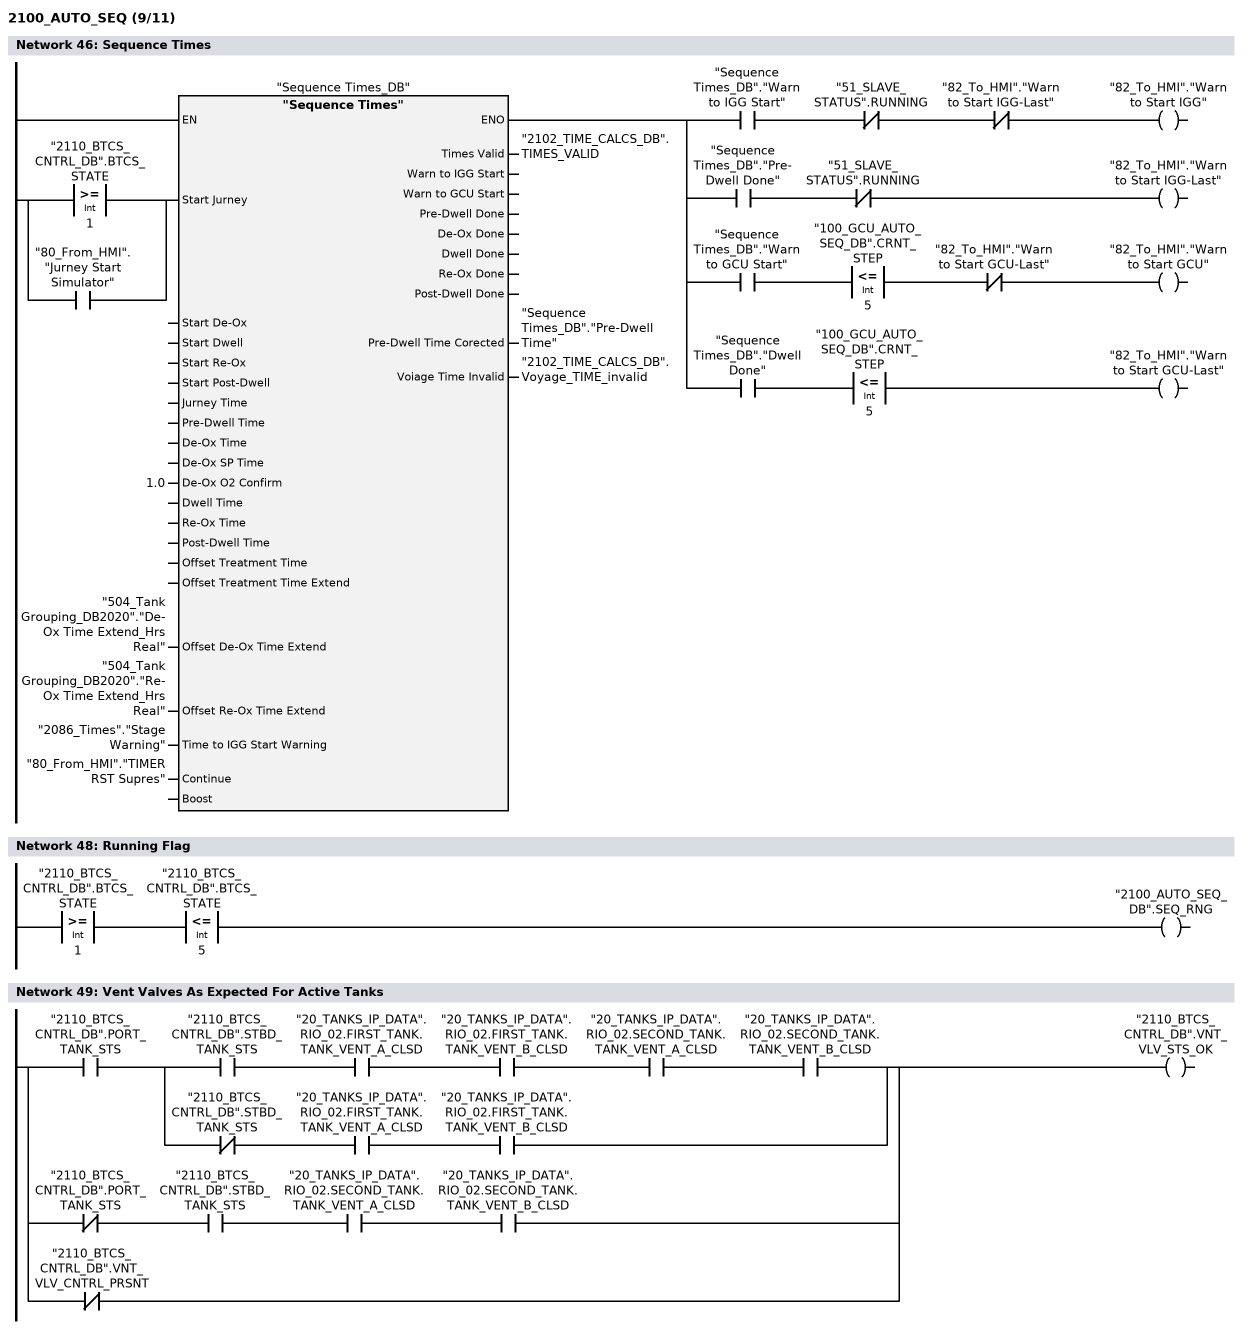
   RUNG wire#powerrail
      "Sequence Times_DB"("Start Jurney" := wire#w1, "Start De-Ox" :=, "Start Dwell" :=, "Start Re-Ox" :=, "Start Post-Dwell" :=, "Jurney Time" :=, "Pre-Dwell Time" :=, "De-Ox Time" :=, "De-Ox SP Time" :=, "De-Ox O2 Confirm" := 1.0, "Dwell Time" :=, "Re-Ox Time" :=, "Post-Dwell Time" :=, "Offset Treatment Time" :=, "Offset Treatment Time Extend" :=, "Offset De-Ox Time Extend" := "504_Tank Grouping_DB2020"."De-Ox Time Extend_Hrs Real", "Offset Re-Ox Time Extend" := "504_Tank Grouping_DB2020"."Re-Ox Time Extend_Hrs Real", "Time to IGG Start Warning" := "2086_Times"."Stage Warning", Continue := "80_From_HMI"."TIMER RST Supres", Boost :=, "Times Valid" => "2102_TIME_CALCS_DB".TIMES_VALID, "Warn to IGG Start" =>, "Warn to GCU Start" =>, "Pre-Dwell Done" =>, "De-Ox Done" =>, "Dwell Done" =>, "Re-Ox Done" =>, "Post-Dwell Done" =>, "Pre-Dwell Time Corected" => "Sequence Times_DB"."Pre-Dwell Time", "Voiage Time Invalid" => "2102_TIME_CALCS_DB".Voyage_TIME_invalid)
      wire#w2
      Contact( "Sequence Times_DB"."Warn to IGG Start" )
      I_Contact( "51_SLAVE_STATUS".RUNNING )
      I_Contact( "82_To_HMI"."Warn to Start IGG-Last" )
      Coil( "82_To_HMI"."Warn to Start IGG" )
   END_RUNG
   RUNG wire#powerrail
      { S7_Templates := "SrcType := Int" } GE_Contact(in1 := "2110_BTCS_CNTRL_DB".BTCS_STATE, in2 := 1)
   END_RUNG wire#w1
   RUNG wire#powerrail
      Contact( "80_From_HMI"."Jurney Start Simulator" )
   END_RUNG wire#w1
   RUNG wire#w2
      Contact( "Sequence Times_DB"."Pre-Dwell Done" )
      I_Contact( "51_SLAVE_STATUS".RUNNING )
      Coil( "82_To_HMI"."Warn to Start IGG-Last" )
   END_RUNG
   RUNG wire#w2
      Contact( "Sequence Times_DB"."Warn to GCU Start" )
      { S7_Templates := "SrcType := Int" } LE_Contact(in1 := "100_GCU_AUTO_SEQ_DB".CRNT_STEP, in2 := 5)
      I_Contact( "82_To_HMI"."Warn to Start GCU-Last" )
      Coil( "82_To_HMI"."Warn to Start GCU" )
   END_RUNG
   RUNG wire#w2
      Contact( "Sequence Times_DB"."Dwell Done" )
      { S7_Templates := "SrcType := Int" } LE_Contact(in1 := "100_GCU_AUTO_SEQ_DB".CRNT_STEP, in2 := 5)
      Coil( "82_To_HMI"."Warn to Start GCU-Last" )
   END_RUNG
   // the same network as SCL:
   "Sequence Times_DB"("Start Jurney" := ("2110_BTCS_CNTRL_DB".BTCS_STATE >= 1) OR "80_From_HMI"."Jurney Start Simulator",   // "Sequence Times"
                       "De-Ox O2 Confirm" := 1.0,
                       "Offset De-Ox Time Extend" := "504_Tank Grouping_DB2020"."De-Ox Time Extend_Hrs Real",
                       "Offset Re-Ox Time Extend" := "504_Tank Grouping_DB2020"."Re-Ox Time Extend_Hrs Real",
                       "Time to IGG Start Warning" := "2086_Times"."Stage Warning",
                       Continue := "80_From_HMI"."TIMER RST Supres",
                       "Times Valid" => "2102_TIME_CALCS_DB".TIMES_VALID,
                       "Pre-Dwell Time Corected" => "Sequence Times_DB"."Pre-Dwell Time",
                       "Voiage Time Invalid" => "2102_TIME_CALCS_DB".Voyage_TIME_invalid,
                       ENO => #_w1);
   "82_To_HMI"."Warn to Start IGG" := #_w1 AND "Sequence Times_DB"."Warn to IGG Start" AND NOT "51_SLAVE_STATUS".RUNNING AND NOT "82_To_HMI"."Warn to Start IGG-Last";
   "82_To_HMI"."Warn to Start IGG-Last" := #_w1 AND "Sequence Times_DB"."Pre-Dwell Done" AND NOT "51_SLAVE_STATUS".RUNNING;
   "82_To_HMI"."Warn to Start GCU" := #_w1 AND "Sequence Times_DB"."Warn to GCU Start" AND ("100_GCU_AUTO_SEQ_DB".CRNT_STEP <= 5) AND NOT "82_To_HMI"."Warn to Start GCU-Last";
   "82_To_HMI"."Warn to Start GCU-Last" := #_w1 AND "Sequence Times_DB"."Dwell Done" AND ("100_GCU_AUTO_SEQ_DB".CRNT_STEP <= 5);
END_REGION

REGION Network 48: Running Flag
   RUNG wire#powerrail
      { S7_Templates := "SrcType := Int" } GE_Contact(in1 := "2110_BTCS_CNTRL_DB".BTCS_STATE, in2 := 1)
      { S7_Templates := "SrcType := Int" } LE_Contact(in1 := "2110_BTCS_CNTRL_DB".BTCS_STATE, in2 := 5)
      Coil( "2100_AUTO_SEQ_DB".SEQ_RNG )
   END_RUNG
   // the same network as SCL:
   "2100_AUTO_SEQ_DB".SEQ_RNG := ("2110_BTCS_CNTRL_DB".BTCS_STATE >= 1) AND ("2110_BTCS_CNTRL_DB".BTCS_STATE <= 5);
END_REGION

REGION Network 49: Vent Valves As Expected For Active Tanks
   RUNG wire#powerrail
      Contact( "2110_BTCS_CNTRL_DB".PORT_TANK_STS )
      wire#w1
      Contact( "2110_BTCS_CNTRL_DB".STBD_TANK_STS )
      Contact( "20_TANKS_IP_DATA".RIO_02.FIRST_TANK.TANK_VENT_A_CLSD )
      Contact( "20_TANKS_IP_DATA".RIO_02.FIRST_TANK.TANK_VENT_B_CLSD )
      Contact( "20_TANKS_IP_DATA".RIO_02.SECOND_TANK.TANK_VENT_A_CLSD )
      Contact( "20_TANKS_IP_DATA".RIO_02.SECOND_TANK.TANK_VENT_B_CLSD )
      wire#w2
      Coil( "2110_BTCS_CNTRL_DB".VNT_VLV_STS_OK )
   END_RUNG
   RUNG wire#w1
      I_Contact( "2110_BTCS_CNTRL_DB".STBD_TANK_STS )
      Contact( "20_TANKS_IP_DATA".RIO_02.FIRST_TANK.TANK_VENT_A_CLSD )
      Contact( "20_TANKS_IP_DATA".RIO_02.FIRST_TANK.TANK_VENT_B_CLSD )
   END_RUNG wire#w2
   RUNG wire#powerrail
      I_Contact( "2110_BTCS_CNTRL_DB".PORT_TANK_STS )
      Contact( "2110_BTCS_CNTRL_DB".STBD_TANK_STS )
      Contact( "20_TANKS_IP_DATA".RIO_02.SECOND_TANK.TANK_VENT_A_CLSD )
      Contact( "20_TANKS_IP_DATA".RIO_02.SECOND_TANK.TANK_VENT_B_CLSD )
   END_RUNG wire#w2
   RUNG wire#powerrail
      I_Contact( "2110_BTCS_CNTRL_DB".VNT_VLV_CNTRL_PRSNT )
   END_RUNG wire#w2
   // the same network as SCL:
   "2110_BTCS_CNTRL_DB".VNT_VLV_STS_OK := ("2110_BTCS_CNTRL_DB".PORT_TANK_STS AND (("2110_BTCS_CNTRL_DB".STBD_TANK_STS AND "20_TANKS_IP_DATA".RIO_02.FIRST_TANK.TANK_VENT_A_CLSD AND "20_TANKS_IP_DATA".RIO_02.FIRST_TANK.TANK_VENT_B_CLSD AND "20_TANKS_IP_DATA".RIO_02.SECOND_TANK.TANK_VENT_A_CLSD AND "20_TANKS_IP_DATA".RIO_02.SECOND_TANK.TANK_VENT_B_CLSD) OR (NOT "2110_BTCS_CNTRL_DB".STBD_TANK_STS AND "20_TANKS_IP_DATA".RIO_02.FIRST_TANK.TANK_VENT_A_CLSD AND "20_TANKS_IP_DATA".RIO_02.FIRST_TANK.TANK_VENT_B_CLSD))) OR (NOT "2110_BTCS_CNTRL_DB".PORT_TANK_STS AND "2110_BTCS_CNTRL_DB".STBD_TANK_STS AND "20_TANKS_IP_DATA".RIO_02.SECOND_TANK.TANK_VENT_A_CLSD AND "20_TANKS_IP_DATA".RIO_02.SECOND_TANK.TANK_VENT_B_CLSD) OR NOT "2110_BTCS_CNTRL_DB".VNT_VLV_CNTRL_PRSNT;
END_REGION

REGION Network 50: GTT Valves As Expected For Active Tanks (condition used from Tank Grouping FB)
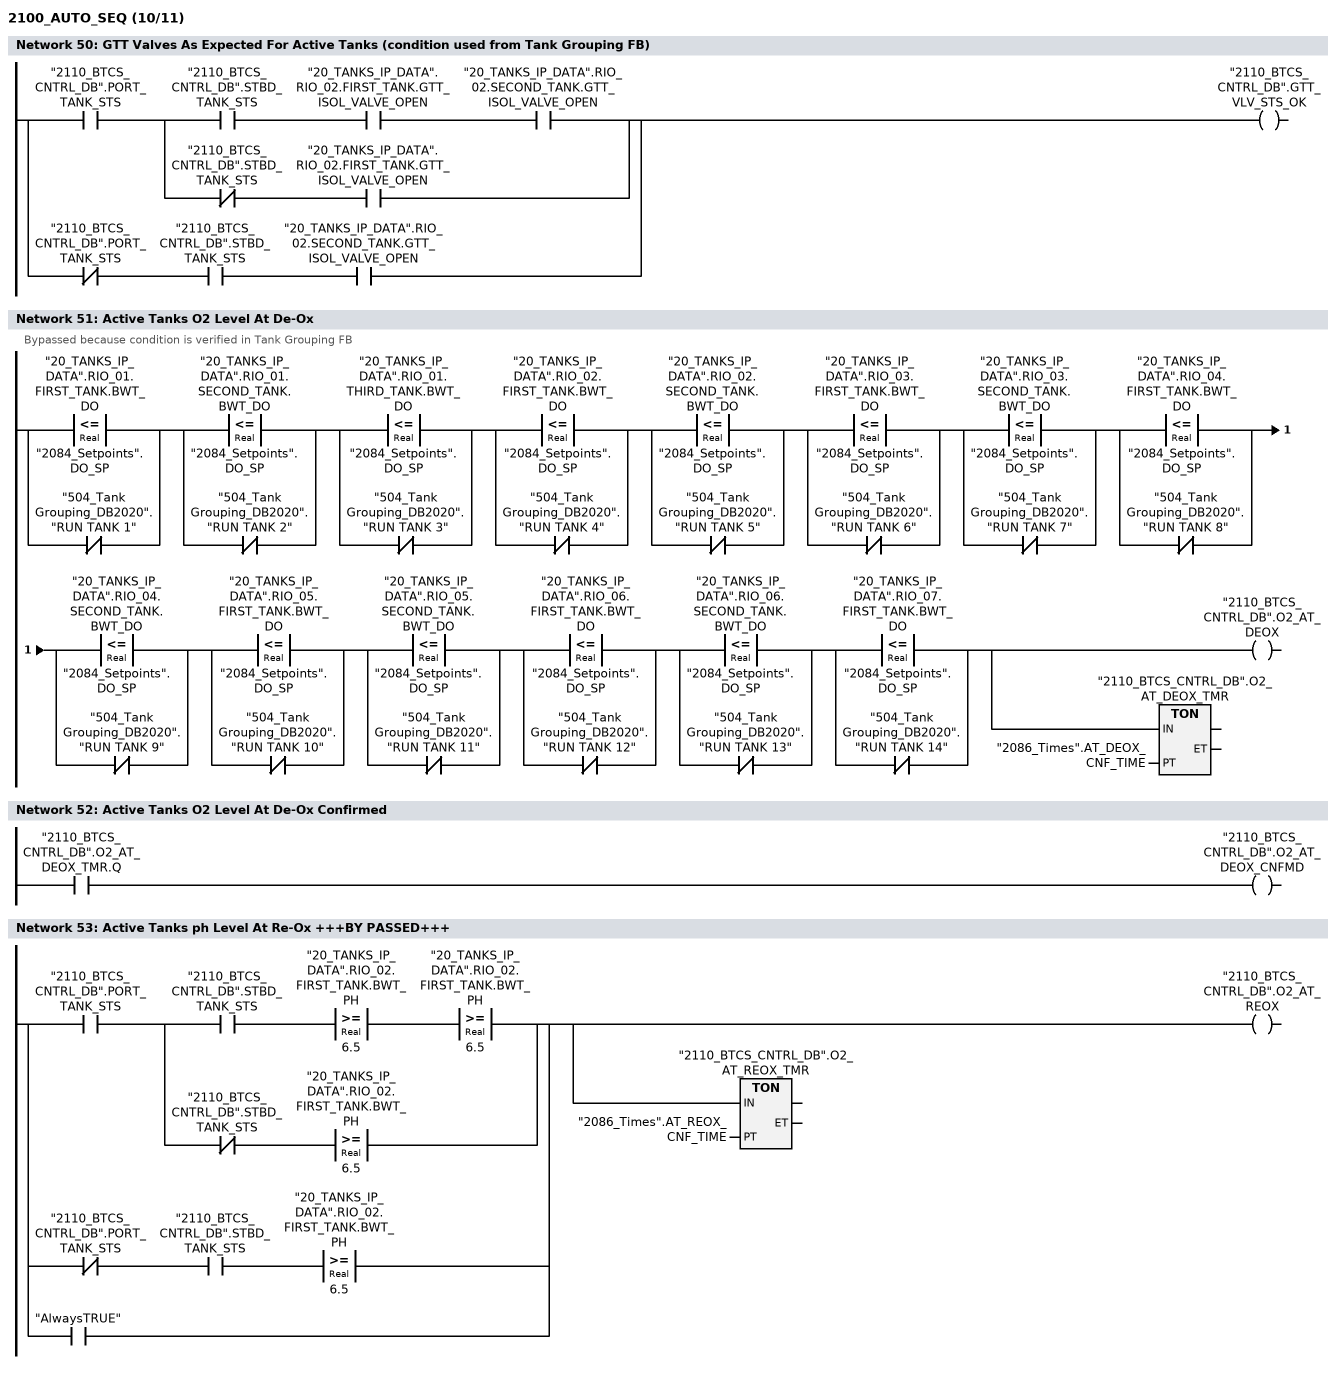
   RUNG wire#powerrail
      Contact( "2110_BTCS_CNTRL_DB".PORT_TANK_STS )
      wire#w1
      Contact( "2110_BTCS_CNTRL_DB".STBD_TANK_STS )
      Contact( "20_TANKS_IP_DATA".RIO_02.FIRST_TANK.GTT_ISOL_VALVE_OPEN )
      Contact( "20_TANKS_IP_DATA".RIO_02.SECOND_TANK.GTT_ISOL_VALVE_OPEN )
      wire#w2
      Coil( "2110_BTCS_CNTRL_DB".GTT_VLV_STS_OK )
   END_RUNG
   RUNG wire#w1
      I_Contact( "2110_BTCS_CNTRL_DB".STBD_TANK_STS )
      Contact( "20_TANKS_IP_DATA".RIO_02.FIRST_TANK.GTT_ISOL_VALVE_OPEN )
   END_RUNG wire#w2
   RUNG wire#powerrail
      I_Contact( "2110_BTCS_CNTRL_DB".PORT_TANK_STS )
      Contact( "2110_BTCS_CNTRL_DB".STBD_TANK_STS )
      Contact( "20_TANKS_IP_DATA".RIO_02.SECOND_TANK.GTT_ISOL_VALVE_OPEN )
   END_RUNG wire#w2
   // the same network as SCL:
   "2110_BTCS_CNTRL_DB".GTT_VLV_STS_OK := ("2110_BTCS_CNTRL_DB".PORT_TANK_STS AND (("2110_BTCS_CNTRL_DB".STBD_TANK_STS AND "20_TANKS_IP_DATA".RIO_02.FIRST_TANK.GTT_ISOL_VALVE_OPEN AND "20_TANKS_IP_DATA".RIO_02.SECOND_TANK.GTT_ISOL_VALVE_OPEN) OR (NOT "2110_BTCS_CNTRL_DB".STBD_TANK_STS AND "20_TANKS_IP_DATA".RIO_02.FIRST_TANK.GTT_ISOL_VALVE_OPEN))) OR (NOT "2110_BTCS_CNTRL_DB".PORT_TANK_STS AND "2110_BTCS_CNTRL_DB".STBD_TANK_STS AND "20_TANKS_IP_DATA".RIO_02.SECOND_TANK.GTT_ISOL_VALVE_OPEN);
END_REGION

REGION Network 51: Active Tanks O2 Level At De-Ox
   // Bypassed because condition is verified in Tank Grouping FB
   "2110_BTCS_CNTRL_DB".O2_AT_DEOX := (("20_TANKS_IP_DATA".RIO_01.FIRST_TANK.BWT_DO <= "2084_Setpoints".DO_SP) OR NOT "504_Tank Grouping_DB2020"."RUN TANK 1") AND (("20_TANKS_IP_DATA".RIO_01.SECOND_TANK.BWT_DO <= "2084_Setpoints".DO_SP) OR NOT "504_Tank Grouping_DB2020"."RUN TANK 2") AND (("20_TANKS_IP_DATA".RIO_01.THIRD_TANK.BWT_DO <= "2084_Setpoints".DO_SP) OR NOT "504_Tank Grouping_DB2020"."RUN TANK 3") AND (("20_TANKS_IP_DATA".RIO_02.FIRST_TANK.BWT_DO <= "2084_Setpoints".DO_SP) OR NOT "504_Tank Grouping_DB2020"."RUN TANK 4") AND (("20_TANKS_IP_DATA".RIO_02.SECOND_TANK.BWT_DO <= "2084_Setpoints".DO_SP) OR NOT "504_Tank Grouping_DB2020"."RUN TANK 5") AND (("20_TANKS_IP_DATA".RIO_03.FIRST_TANK.BWT_DO <= "2084_Setpoints".DO_SP) OR NOT "504_Tank Grouping_DB2020"."RUN TANK 6") AND (("20_TANKS_IP_DATA".RIO_03.SECOND_TANK.BWT_DO <= "2084_Setpoints".DO_SP) OR NOT "504_Tank Grouping_DB2020"."RUN TANK 7") AND (("20_TANKS_IP_DATA".RIO_04.FIRST_TANK.BWT_DO <= "2084_Setpoints".DO_SP) OR NOT "504_Tank Grouping_DB2020"."RUN TANK 8") AND (("20_TANKS_IP_DATA".RIO_04.SECOND_TANK.BWT_DO <= "2084_Setpoints".DO_SP) OR NOT "504_Tank Grouping_DB2020"."RUN TANK 9") AND (("20_TANKS_IP_DATA".RIO_05.FIRST_TANK.BWT_DO <= "2084_Setpoints".DO_SP) OR NOT "504_Tank Grouping_DB2020"."RUN TANK 10") AND (("20_TANKS_IP_DATA".RIO_05.SECOND_TANK.BWT_DO <= "2084_Setpoints".DO_SP) OR NOT "504_Tank Grouping_DB2020"."RUN TANK 11") AND (("20_TANKS_IP_DATA".RIO_06.FIRST_TANK.BWT_DO <= "2084_Setpoints".DO_SP) OR NOT "504_Tank Grouping_DB2020"."RUN TANK 12") AND (("20_TANKS_IP_DATA".RIO_06.SECOND_TANK.BWT_DO <= "2084_Setpoints".DO_SP) OR NOT "504_Tank Grouping_DB2020"."RUN TANK 13") AND (("20_TANKS_IP_DATA".RIO_07.FIRST_TANK.BWT_DO <= "2084_Setpoints".DO_SP) OR NOT "504_Tank Grouping_DB2020"."RUN TANK 14");
   "2110_BTCS_CNTRL_DB".O2_AT_DEOX_TMR.TON(IN := "2110_BTCS_CNTRL_DB".O2_AT_DEOX,
                           PT := "2086_Times".AT_DEOX_CNF_TIME);
END_REGION

REGION Network 52: Active Tanks O2 Level At De-Ox Confirmed
   RUNG wire#powerrail
      Contact( "2110_BTCS_CNTRL_DB".O2_AT_DEOX_TMR.Q )
      Coil( "2110_BTCS_CNTRL_DB".O2_AT_DEOX_CNFMD )
   END_RUNG
   // the same network as SCL:
   "2110_BTCS_CNTRL_DB".O2_AT_DEOX_CNFMD := "2110_BTCS_CNTRL_DB".O2_AT_DEOX_TMR.Q;
END_REGION

REGION Network 53: Active Tanks ph Level At Re-Ox +++BY PASSED+++
   "2110_BTCS_CNTRL_DB".O2_AT_REOX := ("2110_BTCS_CNTRL_DB".PORT_TANK_STS AND (("2110_BTCS_CNTRL_DB".STBD_TANK_STS AND ("20_TANKS_IP_DATA".RIO_02.FIRST_TANK.BWT_PH >= 6.5) AND ("20_TANKS_IP_DATA".RIO_02.FIRST_TANK.BWT_PH >= 6.5)) OR (NOT "2110_BTCS_CNTRL_DB".STBD_TANK_STS AND ("20_TANKS_IP_DATA".RIO_02.FIRST_TANK.BWT_PH >= 6.5)))) OR (NOT "2110_BTCS_CNTRL_DB".PORT_TANK_STS AND "2110_BTCS_CNTRL_DB".STBD_TANK_STS AND ("20_TANKS_IP_DATA".RIO_02.FIRST_TANK.BWT_PH >= 6.5)) OR "AlwaysTRUE";
   "2110_BTCS_CNTRL_DB".O2_AT_REOX_TMR.TON(IN := "2110_BTCS_CNTRL_DB".O2_AT_REOX,
                           PT := "2086_Times".AT_REOX_CNF_TIME);
END_REGION

REGION Network 54: Active Tanks ph Level At Re-Ox Confirmed
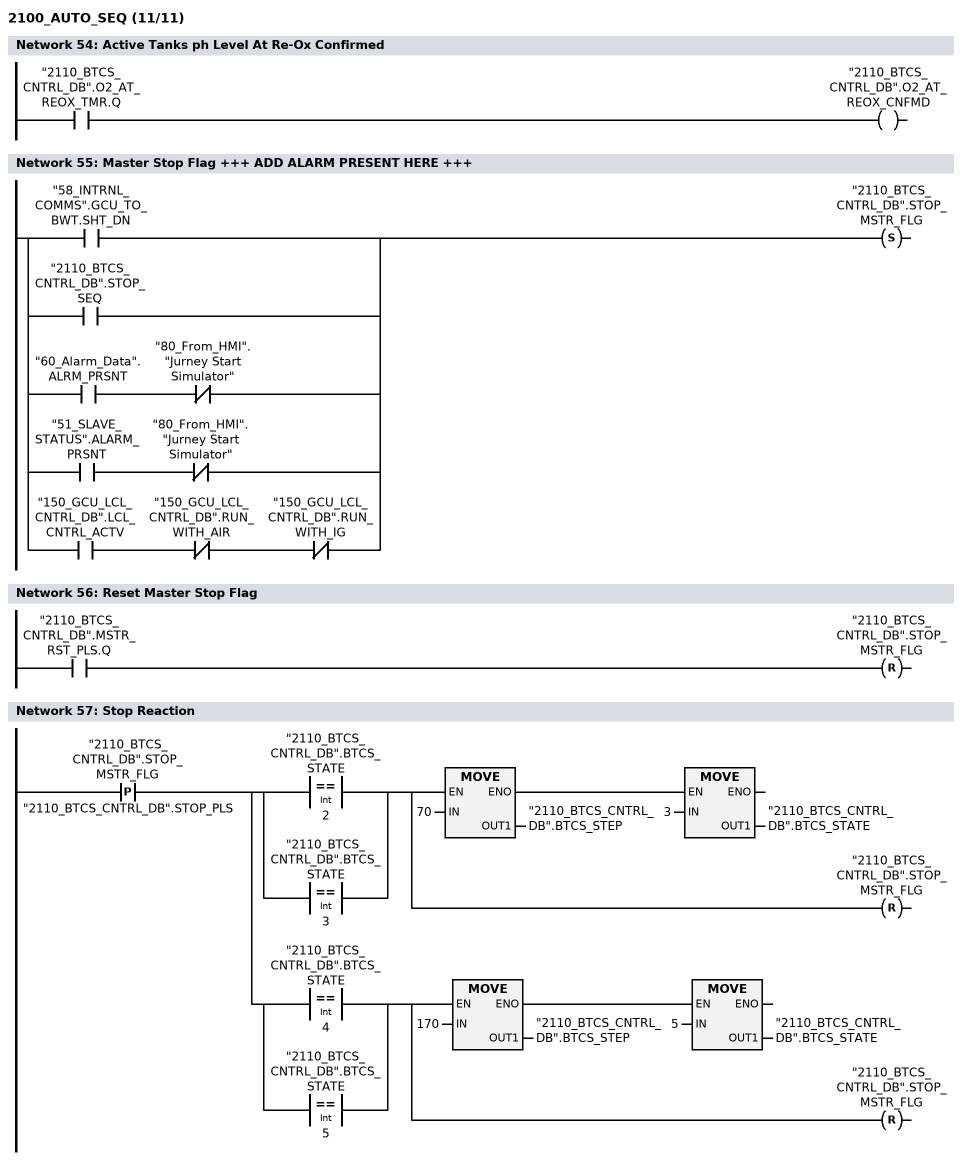
   RUNG wire#powerrail
      Contact( "2110_BTCS_CNTRL_DB".O2_AT_REOX_TMR.Q )
      Coil( "2110_BTCS_CNTRL_DB".O2_AT_REOX_CNFMD )
   END_RUNG
   // the same network as SCL:
   "2110_BTCS_CNTRL_DB".O2_AT_REOX_CNFMD := "2110_BTCS_CNTRL_DB".O2_AT_REOX_TMR.Q;
END_REGION

REGION Network 55: Master Stop Flag +++ ADD ALARM PRESENT HERE +++
   RUNG wire#powerrail
      Contact( "58_INTRNL_COMMS".GCU_TO_BWT.SHT_DN )
      wire#w1
      S_Coil( "2110_BTCS_CNTRL_DB".STOP_MSTR_FLG )
   END_RUNG
   RUNG wire#powerrail
      Contact( "2110_BTCS_CNTRL_DB".STOP_SEQ )
   END_RUNG wire#w1
   RUNG wire#powerrail
      Contact( "60_Alarm_Data".ALRM_PRSNT )
      I_Contact( "80_From_HMI"."Jurney Start Simulator" )
   END_RUNG wire#w1
   RUNG wire#powerrail
      Contact( "51_SLAVE_STATUS".ALARM_PRSNT )
      I_Contact( "80_From_HMI"."Jurney Start Simulator" )
   END_RUNG wire#w1
   RUNG wire#powerrail
      Contact( "150_GCU_LCL_CNTRL_DB".LCL_CNTRL_ACTV )
      I_Contact( "150_GCU_LCL_CNTRL_DB".RUN_WITH_AIR )
      I_Contact( "150_GCU_LCL_CNTRL_DB".RUN_WITH_IG )
   END_RUNG wire#w1
   // the same network as SCL:
   IF "58_INTRNL_COMMS".GCU_TO_BWT.SHT_DN OR "2110_BTCS_CNTRL_DB".STOP_SEQ OR ("60_Alarm_Data".ALRM_PRSNT AND NOT "80_From_HMI"."Jurney Start Simulator") OR ("51_SLAVE_STATUS".ALARM_PRSNT AND NOT "80_From_HMI"."Jurney Start Simulator") OR ("150_GCU_LCL_CNTRL_DB".LCL_CNTRL_ACTV AND NOT "150_GCU_LCL_CNTRL_DB".RUN_WITH_AIR AND NOT "150_GCU_LCL_CNTRL_DB".RUN_WITH_IG) THEN
       "2110_BTCS_CNTRL_DB".STOP_MSTR_FLG := TRUE;
   END_IF;
END_REGION

REGION Network 56: Reset Master Stop Flag
   RUNG wire#powerrail
      Contact( "2110_BTCS_CNTRL_DB".MSTR_RST_PLS.Q )
      R_Coil( "2110_BTCS_CNTRL_DB".STOP_MSTR_FLG )
   END_RUNG
   // the same network as SCL:
   IF "2110_BTCS_CNTRL_DB".MSTR_RST_PLS.Q THEN "2110_BTCS_CNTRL_DB".STOP_MSTR_FLG := FALSE; END_IF;
END_REGION

REGION Network 57: Stop Reaction
   RUNG wire#powerrail
      P_Contact(operand := "2110_BTCS_CNTRL_DB".STOP_MSTR_FLG, bit := "2110_BTCS_CNTRL_DB".STOP_PLS)
      wire#w1
      { S7_Templates := "SrcType := Int" } EQ_Contact(in1 := "2110_BTCS_CNTRL_DB".BTCS_STATE, in2 := 2)
      wire#w2
      Move(in := 70, out1 => "2110_BTCS_CNTRL_DB".BTCS_STEP)
      Move(in := 3, out1 => "2110_BTCS_CNTRL_DB".BTCS_STATE)
   END_RUNG
   RUNG wire#w1
      { S7_Templates := "SrcType := Int" } EQ_Contact(in1 := "2110_BTCS_CNTRL_DB".BTCS_STATE, in2 := 3)
   END_RUNG wire#w2
   RUNG wire#w2
      R_Coil( "2110_BTCS_CNTRL_DB".STOP_MSTR_FLG )
   END_RUNG
   RUNG wire#w1
      { S7_Templates := "SrcType := Int" } EQ_Contact(in1 := "2110_BTCS_CNTRL_DB".BTCS_STATE, in2 := 4)
      wire#w3
      Move(in := 170, out1 => "2110_BTCS_CNTRL_DB".BTCS_STEP)
      Move(in := 5, out1 => "2110_BTCS_CNTRL_DB".BTCS_STATE)
   END_RUNG
   RUNG wire#w1
      { S7_Templates := "SrcType := Int" } EQ_Contact(in1 := "2110_BTCS_CNTRL_DB".BTCS_STATE, in2 := 5)
   END_RUNG wire#w3
   RUNG wire#w3
      R_Coil( "2110_BTCS_CNTRL_DB".STOP_MSTR_FLG )
   END_RUNG
   // the same network as SCL:
   #_w1 := "2110_BTCS_CNTRL_DB".STOP_MSTR_FLG AND NOT "2110_BTCS_CNTRL_DB".STOP_PLS;   // rising edge of "2110_BTCS_CNTRL_DB".STOP_MSTR_FLG
   "2110_BTCS_CNTRL_DB".STOP_PLS := "2110_BTCS_CNTRL_DB".STOP_MSTR_FLG;
   IF #_w1 AND (("2110_BTCS_CNTRL_DB".BTCS_STATE = 2) OR ("2110_BTCS_CNTRL_DB".BTCS_STATE = 3)) THEN
       "2110_BTCS_CNTRL_DB".BTCS_STEP := 70;
   END_IF;
   #_w2 := #_w1 AND (("2110_BTCS_CNTRL_DB".BTCS_STATE = 2) OR ("2110_BTCS_CNTRL_DB".BTCS_STATE = 3));
   IF #_w2 THEN
       "2110_BTCS_CNTRL_DB".BTCS_STATE := 3;
       "2110_BTCS_CNTRL_DB".STOP_MSTR_FLG := FALSE;
   END_IF;
   IF #_w1 AND (("2110_BTCS_CNTRL_DB".BTCS_STATE = 4) OR ("2110_BTCS_CNTRL_DB".BTCS_STATE = 5)) THEN
       "2110_BTCS_CNTRL_DB".BTCS_STEP := 170;
   END_IF;
   #_w3 := #_w1 AND (("2110_BTCS_CNTRL_DB".BTCS_STATE = 4) OR ("2110_BTCS_CNTRL_DB".BTCS_STATE = 5));
   IF #_w3 THEN
       "2110_BTCS_CNTRL_DB".BTCS_STATE := 5;
       "2110_BTCS_CNTRL_DB".STOP_MSTR_FLG := FALSE;
   END_IF;
END_REGION
END_FUNCTION

FUNCTION "2102_TIME_CALCS" : Void   // FC2102, LAD
TITLE = Time Calculations
{ S7_Optimized_Access := 'TRUE' }
AUTHOR : JRS
VERSION : 0.1
// For calculating time periods associated with the BTCS
   VAR_TEMP
      T_REAL : Real;
   END_VAR
   VAR_TEMP   // added for the SCL form of the ladder/FBD networks
      _w1 : Bool;
      _w2 : Bool;
      _w3 : Bool;
      _w4 : Bool;
      _w5 : Bool;
      _w6 : Bool;
      _w7 : Bool;
   END_VAR
BEGIN

REGION Network 2: Minutes Phase Difference
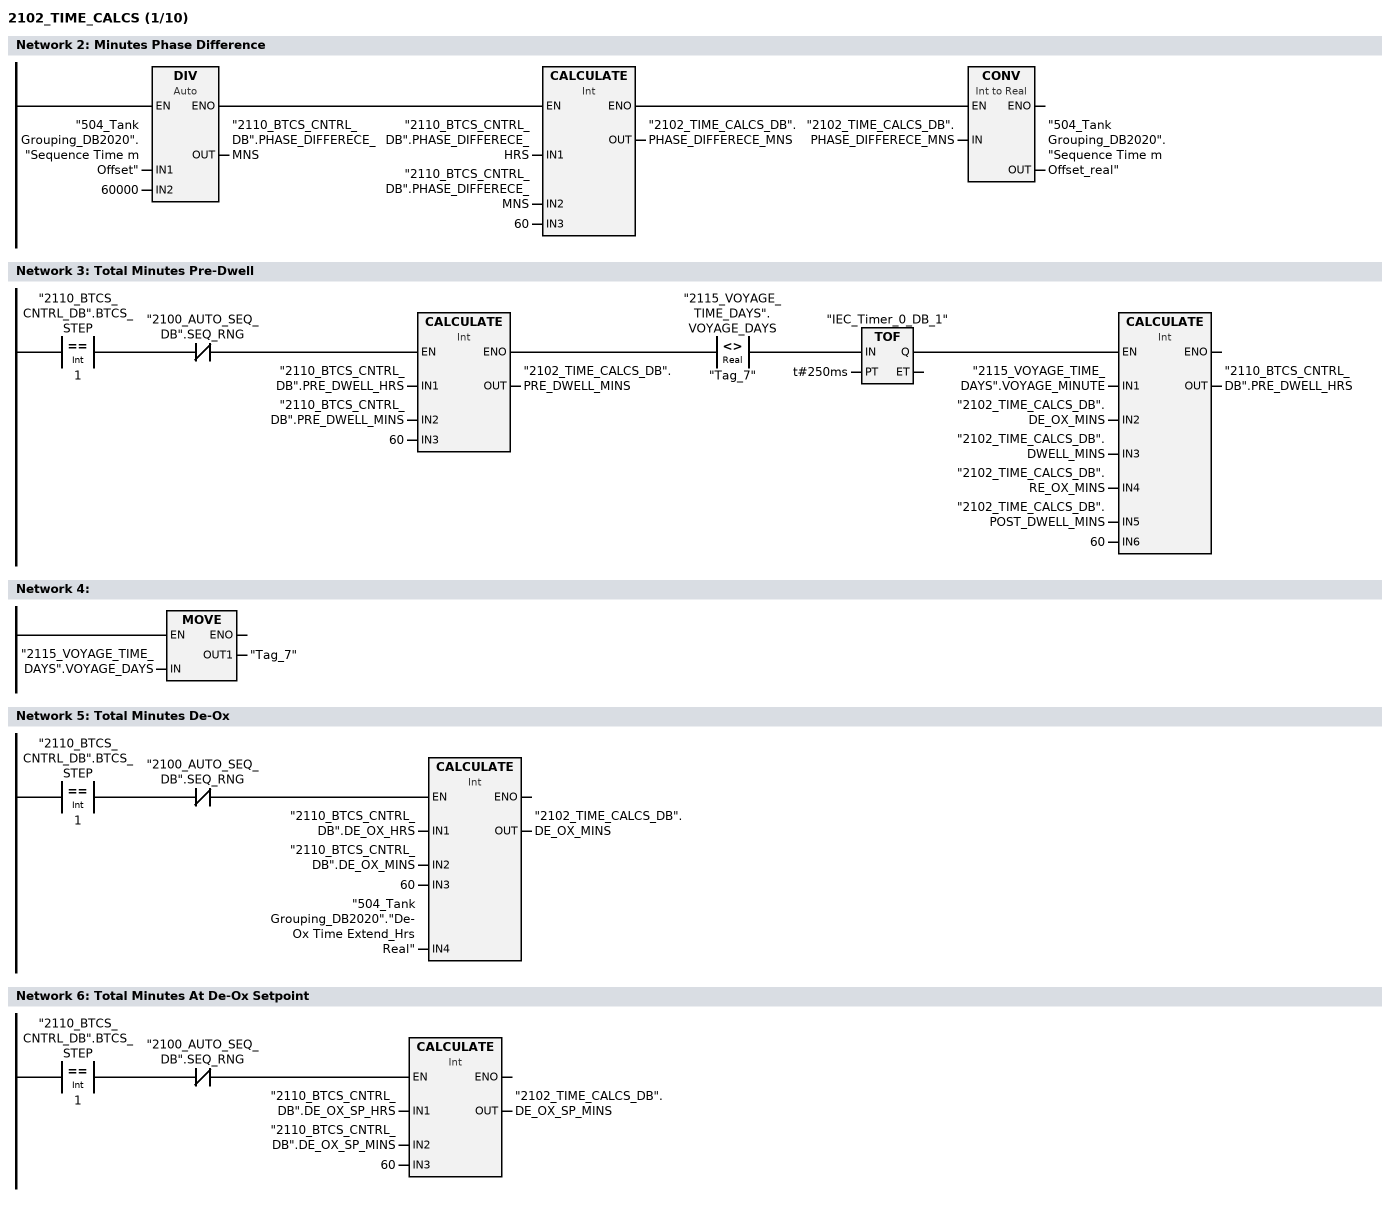
   RUNG wire#powerrail
      Div(in1 := "504_Tank Grouping_DB2020"."Sequence Time m Offset", in2 := 60000, out => "2110_BTCS_CNTRL_DB".PHASE_DIFFERECE_MNS)
      { S7_Templates := "SrcType := Int"; S7_Expression := "(IN1*IN3)+IN2" } Calculate(in1 := "2110_BTCS_CNTRL_DB".PHASE_DIFFERECE_HRS, in2 := "2110_BTCS_CNTRL_DB".PHASE_DIFFERECE_MNS, in3 := 60, out => "2102_TIME_CALCS_DB".PHASE_DIFFERECE_MNS)
      { S7_Templates := "[SrcType := Int, DestType := Real]" } Convert(in := "2102_TIME_CALCS_DB".PHASE_DIFFERECE_MNS, out => "504_Tank Grouping_DB2020"."Sequence Time m Offset_real")
   END_RUNG
   // the same network as SCL:
   "2110_BTCS_CNTRL_DB".PHASE_DIFFERECE_MNS := "504_Tank Grouping_DB2020"."Sequence Time m Offset" / 60000;
   "2102_TIME_CALCS_DB".PHASE_DIFFERECE_MNS := ("2110_BTCS_CNTRL_DB".PHASE_DIFFERECE_HRS*60)+"2110_BTCS_CNTRL_DB".PHASE_DIFFERECE_MNS;
   "504_Tank Grouping_DB2020"."Sequence Time m Offset_real" := INT_TO_REAL("2102_TIME_CALCS_DB".PHASE_DIFFERECE_MNS);
END_REGION

REGION Network 3: Total Minutes Pre-Dwell
   #_w1 := ("2110_BTCS_CNTRL_DB".BTCS_STEP = 1) AND NOT "2100_AUTO_SEQ_DB".SEQ_RNG;
   IF #_w1 THEN
       "2102_TIME_CALCS_DB".PRE_DWELL_MINS := ("2110_BTCS_CNTRL_DB".PRE_DWELL_HRS*60)+"2110_BTCS_CNTRL_DB".PRE_DWELL_MINS;
   END_IF;
   "IEC_Timer_0_DB_1".TOF(IN := #_w1 AND ("2115_VOYAGE_TIME_DAYS".VOYAGE_DAYS <> "Tag_7"), PT := t#250ms);
   IF "IEC_Timer_0_DB_1".Q THEN
       "2110_BTCS_CNTRL_DB".PRE_DWELL_HRS := ("2115_VOYAGE_TIME_DAYS".VOYAGE_MINUTE-("2102_TIME_CALCS_DB".DE_OX_MINS+"2102_TIME_CALCS_DB".DWELL_MINS+"2102_TIME_CALCS_DB".RE_OX_MINS+"2102_TIME_CALCS_DB".POST_DWELL_MINS))/60;
   END_IF;
END_REGION

REGION Network 4
   RUNG wire#powerrail
      Move(in := "2115_VOYAGE_TIME_DAYS".VOYAGE_DAYS, out1 => "Tag_7")
   END_RUNG
   // the same network as SCL:
   "Tag_7" := "2115_VOYAGE_TIME_DAYS".VOYAGE_DAYS;
END_REGION

REGION Network 5: Total Minutes De-Ox
   RUNG wire#powerrail
      { S7_Templates := "SrcType := Int" } EQ_Contact(in1 := "2110_BTCS_CNTRL_DB".BTCS_STEP, in2 := 1)
      I_Contact( "2100_AUTO_SEQ_DB".SEQ_RNG )
      { S7_Templates := "SrcType := Int"; S7_Expression := "(IN1*IN3)+IN2+IN4" } Calculate(in1 := "2110_BTCS_CNTRL_DB".DE_OX_HRS, in2 := "2110_BTCS_CNTRL_DB".DE_OX_MINS, in3 := 60, in4 := "504_Tank Grouping_DB2020"."De-Ox Time Extend_Hrs Real", out => "2102_TIME_CALCS_DB".DE_OX_MINS)
   END_RUNG
   // the same network as SCL:
   IF ("2110_BTCS_CNTRL_DB".BTCS_STEP = 1) AND NOT "2100_AUTO_SEQ_DB".SEQ_RNG THEN
       "2102_TIME_CALCS_DB".DE_OX_MINS := ("2110_BTCS_CNTRL_DB".DE_OX_HRS*60)+"2110_BTCS_CNTRL_DB".DE_OX_MINS+"504_Tank Grouping_DB2020"."De-Ox Time Extend_Hrs Real";
   END_IF;
END_REGION

REGION Network 6: Total Minutes At De-Ox Setpoint
   RUNG wire#powerrail
      { S7_Templates := "SrcType := Int" } EQ_Contact(in1 := "2110_BTCS_CNTRL_DB".BTCS_STEP, in2 := 1)
      I_Contact( "2100_AUTO_SEQ_DB".SEQ_RNG )
      { S7_Templates := "SrcType := Int"; S7_Expression := "(IN1*IN3)+IN2" } Calculate(in1 := "2110_BTCS_CNTRL_DB".DE_OX_SP_HRS, in2 := "2110_BTCS_CNTRL_DB".DE_OX_SP_MINS, in3 := 60, out => "2102_TIME_CALCS_DB".DE_OX_SP_MINS)
   END_RUNG
   // the same network as SCL:
   IF ("2110_BTCS_CNTRL_DB".BTCS_STEP = 1) AND NOT "2100_AUTO_SEQ_DB".SEQ_RNG THEN
       "2102_TIME_CALCS_DB".DE_OX_SP_MINS := ("2110_BTCS_CNTRL_DB".DE_OX_SP_HRS*60)+"2110_BTCS_CNTRL_DB".DE_OX_SP_MINS;
   END_IF;
END_REGION

REGION Network 7: Total Minutes Dwell
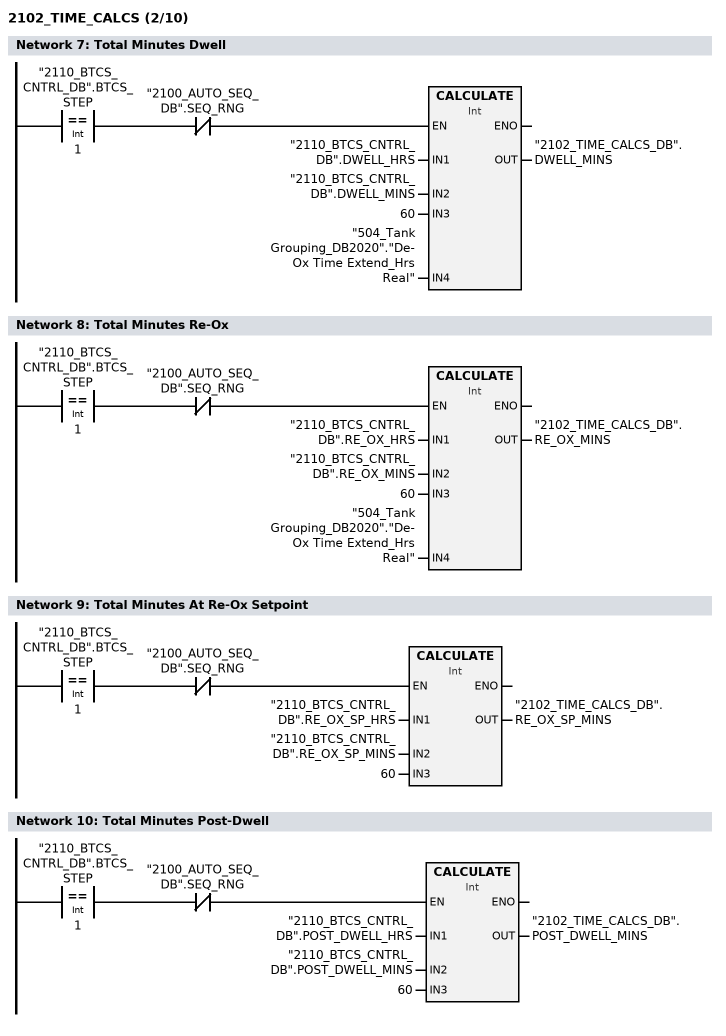
   RUNG wire#powerrail
      { S7_Templates := "SrcType := Int" } EQ_Contact(in1 := "2110_BTCS_CNTRL_DB".BTCS_STEP, in2 := 1)
      I_Contact( "2100_AUTO_SEQ_DB".SEQ_RNG )
      { S7_Templates := "SrcType := Int"; S7_Expression := "(IN1*IN3)+IN2-IN4" } Calculate(in1 := "2110_BTCS_CNTRL_DB".DWELL_HRS, in2 := "2110_BTCS_CNTRL_DB".DWELL_MINS, in3 := 60, in4 := "504_Tank Grouping_DB2020"."De-Ox Time Extend_Hrs Real", out => "2102_TIME_CALCS_DB".DWELL_MINS)
   END_RUNG
   // the same network as SCL:
   IF ("2110_BTCS_CNTRL_DB".BTCS_STEP = 1) AND NOT "2100_AUTO_SEQ_DB".SEQ_RNG THEN
       "2102_TIME_CALCS_DB".DWELL_MINS := ("2110_BTCS_CNTRL_DB".DWELL_HRS*60)+"2110_BTCS_CNTRL_DB".DWELL_MINS-"504_Tank Grouping_DB2020"."De-Ox Time Extend_Hrs Real";
   END_IF;
END_REGION

REGION Network 8: Total Minutes Re-Ox
   RUNG wire#powerrail
      { S7_Templates := "SrcType := Int" } EQ_Contact(in1 := "2110_BTCS_CNTRL_DB".BTCS_STEP, in2 := 1)
      I_Contact( "2100_AUTO_SEQ_DB".SEQ_RNG )
      { S7_Templates := "SrcType := Int"; S7_Expression := "(IN1*IN3)+IN2+IN4" } Calculate(in1 := "2110_BTCS_CNTRL_DB".RE_OX_HRS, in2 := "2110_BTCS_CNTRL_DB".RE_OX_MINS, in3 := 60, in4 := "504_Tank Grouping_DB2020"."De-Ox Time Extend_Hrs Real", out => "2102_TIME_CALCS_DB".RE_OX_MINS)
   END_RUNG
   // the same network as SCL:
   IF ("2110_BTCS_CNTRL_DB".BTCS_STEP = 1) AND NOT "2100_AUTO_SEQ_DB".SEQ_RNG THEN
       "2102_TIME_CALCS_DB".RE_OX_MINS := ("2110_BTCS_CNTRL_DB".RE_OX_HRS*60)+"2110_BTCS_CNTRL_DB".RE_OX_MINS+"504_Tank Grouping_DB2020"."De-Ox Time Extend_Hrs Real";
   END_IF;
END_REGION

REGION Network 9: Total Minutes At Re-Ox Setpoint
   RUNG wire#powerrail
      { S7_Templates := "SrcType := Int" } EQ_Contact(in1 := "2110_BTCS_CNTRL_DB".BTCS_STEP, in2 := 1)
      I_Contact( "2100_AUTO_SEQ_DB".SEQ_RNG )
      { S7_Templates := "SrcType := Int"; S7_Expression := "(IN1*IN3)+IN2" } Calculate(in1 := "2110_BTCS_CNTRL_DB".RE_OX_SP_HRS, in2 := "2110_BTCS_CNTRL_DB".RE_OX_SP_MINS, in3 := 60, out => "2102_TIME_CALCS_DB".RE_OX_SP_MINS)
   END_RUNG
   // the same network as SCL:
   IF ("2110_BTCS_CNTRL_DB".BTCS_STEP = 1) AND NOT "2100_AUTO_SEQ_DB".SEQ_RNG THEN
       "2102_TIME_CALCS_DB".RE_OX_SP_MINS := ("2110_BTCS_CNTRL_DB".RE_OX_SP_HRS*60)+"2110_BTCS_CNTRL_DB".RE_OX_SP_MINS;
   END_IF;
END_REGION

REGION Network 10: Total Minutes Post-Dwell
   RUNG wire#powerrail
      { S7_Templates := "SrcType := Int" } EQ_Contact(in1 := "2110_BTCS_CNTRL_DB".BTCS_STEP, in2 := 1)
      I_Contact( "2100_AUTO_SEQ_DB".SEQ_RNG )
      { S7_Templates := "SrcType := Int"; S7_Expression := "(IN1*IN3)+IN2" } Calculate(in1 := "2110_BTCS_CNTRL_DB".POST_DWELL_HRS, in2 := "2110_BTCS_CNTRL_DB".POST_DWELL_MINS, in3 := 60, out => "2102_TIME_CALCS_DB".POST_DWELL_MINS)
   END_RUNG
   // the same network as SCL:
   IF ("2110_BTCS_CNTRL_DB".BTCS_STEP = 1) AND NOT "2100_AUTO_SEQ_DB".SEQ_RNG THEN
       "2102_TIME_CALCS_DB".POST_DWELL_MINS := ("2110_BTCS_CNTRL_DB".POST_DWELL_HRS*60)+"2110_BTCS_CNTRL_DB".POST_DWELL_MINS;
   END_IF;
END_REGION

REGION Network 11: Total Sequence Time
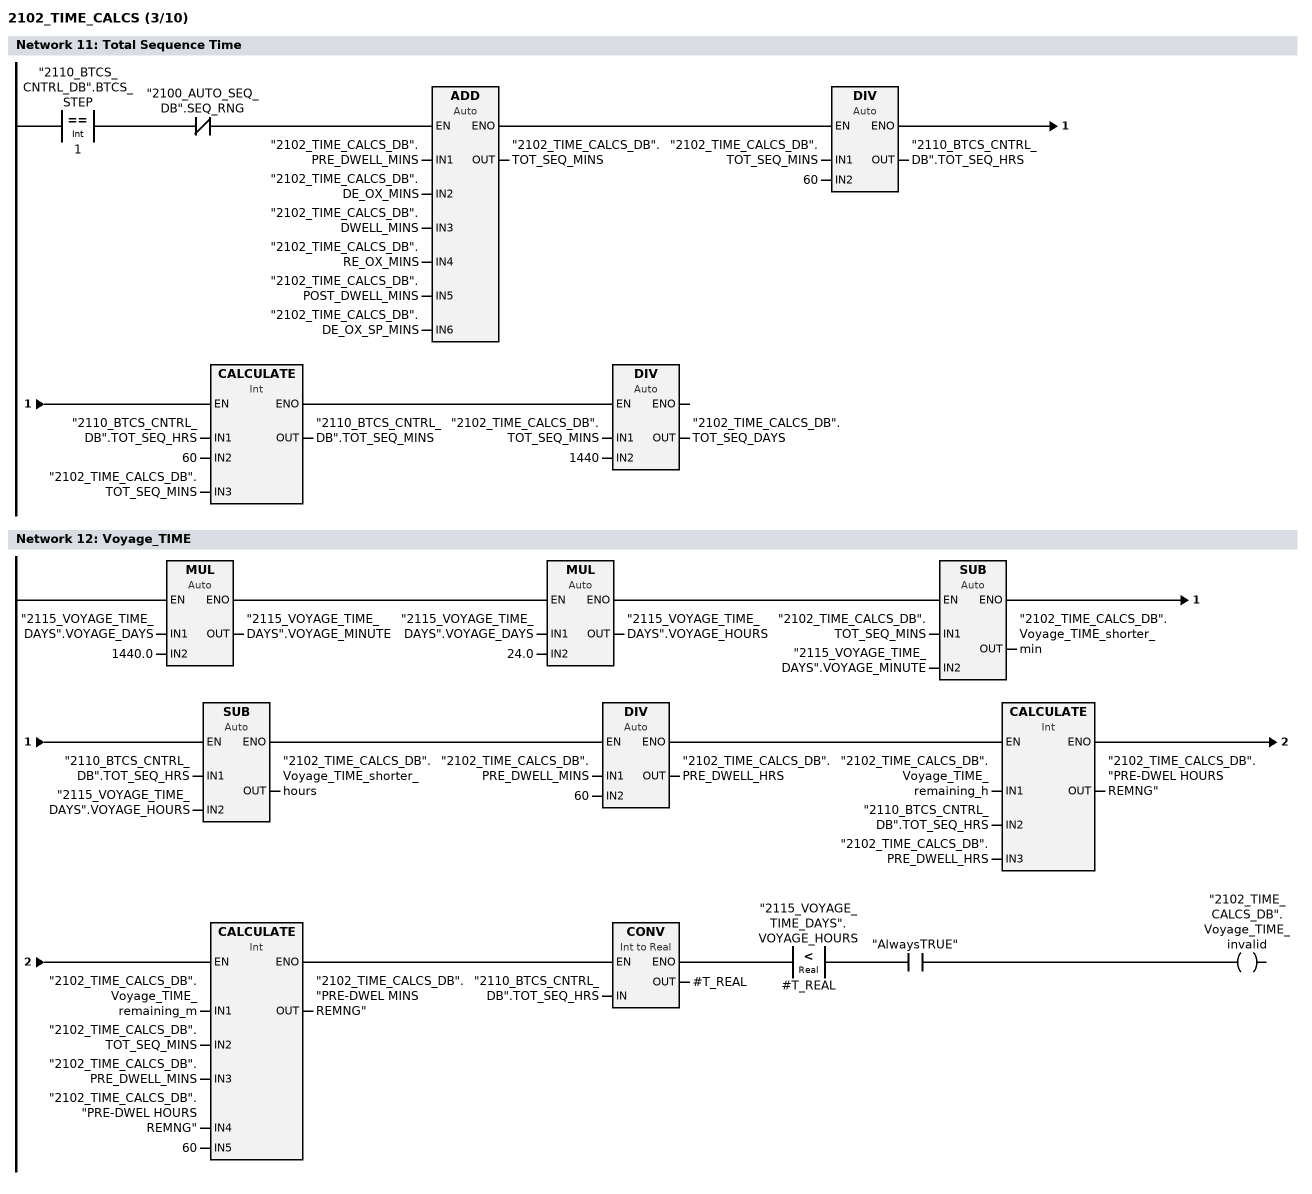
   RUNG wire#powerrail
      { S7_Templates := "SrcType := Int" } EQ_Contact(in1 := "2110_BTCS_CNTRL_DB".BTCS_STEP, in2 := 1)
      I_Contact( "2100_AUTO_SEQ_DB".SEQ_RNG )
      Add(in1 := "2102_TIME_CALCS_DB".PRE_DWELL_MINS, in2 := "2102_TIME_CALCS_DB".DE_OX_MINS, in3 := "2102_TIME_CALCS_DB".DWELL_MINS, in4 := "2102_TIME_CALCS_DB".RE_OX_MINS, in5 := "2102_TIME_CALCS_DB".POST_DWELL_MINS, in6 := "2102_TIME_CALCS_DB".DE_OX_SP_MINS, out => "2102_TIME_CALCS_DB".TOT_SEQ_MINS)
      Div(in1 := "2102_TIME_CALCS_DB".TOT_SEQ_MINS, in2 := 60, out => "2110_BTCS_CNTRL_DB".TOT_SEQ_HRS)
      { S7_Templates := "SrcType := Int"; S7_Expression := "IN3-(IN1*IN2)" } Calculate(in1 := "2110_BTCS_CNTRL_DB".TOT_SEQ_HRS, in2 := 60, in3 := "2102_TIME_CALCS_DB".TOT_SEQ_MINS, out => "2110_BTCS_CNTRL_DB".TOT_SEQ_MINS)
      Div(in1 := "2102_TIME_CALCS_DB".TOT_SEQ_MINS, in2 := 1440, out => "2102_TIME_CALCS_DB".TOT_SEQ_DAYS)
   END_RUNG
   // the same network as SCL:
   IF ("2110_BTCS_CNTRL_DB".BTCS_STEP = 1) AND NOT "2100_AUTO_SEQ_DB".SEQ_RNG THEN
       "2102_TIME_CALCS_DB".TOT_SEQ_MINS := "2102_TIME_CALCS_DB".PRE_DWELL_MINS + "2102_TIME_CALCS_DB".DE_OX_MINS + "2102_TIME_CALCS_DB".DWELL_MINS + "2102_TIME_CALCS_DB".RE_OX_MINS + "2102_TIME_CALCS_DB".POST_DWELL_MINS + "2102_TIME_CALCS_DB".DE_OX_SP_MINS;
       "2110_BTCS_CNTRL_DB".TOT_SEQ_HRS := "2102_TIME_CALCS_DB".TOT_SEQ_MINS / 60;
       "2110_BTCS_CNTRL_DB".TOT_SEQ_MINS := "2102_TIME_CALCS_DB".TOT_SEQ_MINS-("2110_BTCS_CNTRL_DB".TOT_SEQ_HRS*60);
       "2102_TIME_CALCS_DB".TOT_SEQ_DAYS := "2102_TIME_CALCS_DB".TOT_SEQ_MINS / 1440;
   END_IF;
END_REGION
